(* Logix 5000 project; controller FV vendor 1 type 14 code 217 rev 31.11; software revision 31.00; part 43 of 63 *)
(* tags used below, declared in another part *)
   FV_B100 : INT[255];   // FV FLAGS
   FV_F8 : REAL[256];
   FV_FV10C : PlantItem;   // FV10C
   FV_FV10J : PlantItem;   // FV10J
   FV_FV11C : PlantItem;   // FV11C
   FV_FV11J : PlantItem;   // FV11J
   FV_FV12C : PlantItem;   // FV12C
   FV_FV12J : PlantItem;   // FV12J
   FV_FV13C : PlantItem;   // FV13C
   FV_FV13J : PlantItem;   // FV13J
   FV_FV14C : PlantItem;   // FV14C
   FV_FV14J : PlantItem;   // FV14J
   FV_FV15C : PlantItem;   // FV15C
   FV_FV15J : PlantItem;   // FV15J
   FV_FV16C : PlantItem;   // FV16C
   FV_FV16J : PlantItem;   // FV16J
   FV_FV17C : PlantItem;   // FV17C
   FV_FV17J : PlantItem;   // FV17J
   FV_FV18C : PlantItem;   // FV18C
   FV_FV18J : PlantItem;   // FV18J
   FV_FV19C : PlantItem;   // FV19C
   FV_FV19J : PlantItem;   // FV19J
   FV_FV1C : PlantItem;   // FV1C
   FV_FV1J : PlantItem;   // FV1J
   FV_FV20C : PlantItem;   // FV20C
   FV_FV20J : PlantItem;   // FV20J
   FV_FV21C : PlantItem;   // FV21C
   FV_FV21J : PlantItem;   // FV21J
   FV_FV22C : PlantItem;   // FV22C
   FV_FV22J : PlantItem;   // FV22J
   FV_FV2C : PlantItem;   // FV2C
   FV_FV2J : PlantItem;   // FV2J
   FV_FV3C : PlantItem;   // FV3C
   FV_FV3J : PlantItem;   // FV3J
   FV_FV4C : PlantItem;   // FV4C
   FV_FV4J : PlantItem;   // FV4J
   FV_FV5C : PlantItem;   // FV5C
   FV_FV5J : PlantItem;   // FV5J
   FV_FV6C : PlantItem;   // FV6C
   FV_FV6J : PlantItem;   // FV6J
   FV_FV7C : PlantItem;   // FV7C
   FV_FV7J : PlantItem;   // FV7J
   FV_FV8C : PlantItem;   // FV8C
   FV_FV8J : PlantItem;   // FV8J
   FV_FV9C : PlantItem;   // FV9C
   FV_FV9J : PlantItem;   // FV9J
   FV_N101 : INT[255];   // FV INT Fermentation control integer workspace
   FV_N110 : INT[255];   // FV DATA 0 CURRENT FV DATA
   FV_N111 : INT[50];   // FV1, CURRENT FV DATA
   FV_N112 : INT[50];   // FV2, CURRENT FV DATA
   FV_N113 : INT[50];   // FV3, CURRENT FV DATA
   FV_N114 : INT[50];   // FV4, CURRENT FV DATA
   FV_N115 : INT[50];   // FV5, CURRENT FV DATA
   FV_N116 : INT[50];   // FV6, CURRENT FV DATA
   FV_N117 : INT[50];   // FV7, CURRENT FV DATA
   FV_N118 : INT[50];   // FV8, CURRENT FV DATA
   FV_N119 : INT[50];   // FV9, CURRENT FV DATA
   FV_N12 : INT[255];   // SYS_PARMS System Parameter Fil e
   FV_N120 : INT[50];   // FV10, CURRENT FV DATA
   FV_N121 : INT[50];   // FV11, CURRENT FV DATA
   FV_N122 : INT[50];   // FV12, CURRENT FV DATA
   FV_N123 : INT[50];   // FV13, CURRENT FV DATA
   FV_N124 : INT[50];   // FV14, CURRENT FV DATA
   FV_N125 : INT[50];   // FV15, CURRENT FV DATA
   FV_N126 : INT[50];   // FV16, CURRENT FV DATA
   FV_N127 : INT[50];   // FV17, CURRENT FV DATA
   FV_N128 : INT[50];   // FV18, CURRENT FV DATA
   FV_N129 : INT[50];   // FV19, CURRENT FV DATA
   FV_N130 : INT[50];   // FV20, CURRENT FV DATA
   FV_N131 : INT[50];   // FV21, CURRENT FV DATA
   FV_N132 : INT[50];   // FV22, CURRENT FV DATA
   FV_SFile : INT[255];   // SLC Equivalent System File, So Original Code Can Remain
(* FV_Common, continued *)

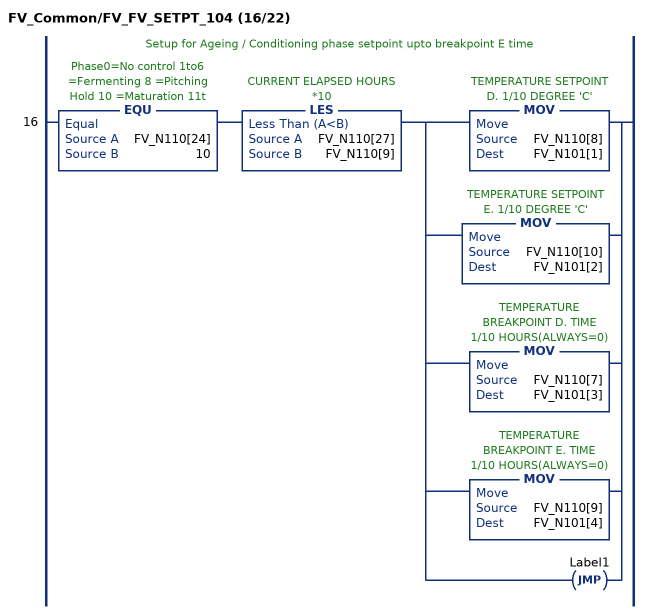
   [picture p920: FV_Common/FV_FV_SETPT_104 rungs 16-16]
   // Setup for Ageing / Conditioning phase setpoint upto breakpoint E time
   16: EQU(FV_N110[24],10)LES(FV_N110[27],FV_N110[9])[MOV(FV_N110[8],FV_N101[1]) ,MOV(FV_N110[10],FV_N101[2]) ,MOV(FV_N110[7],FV_N101[3]) ,MOV(FV_N110[9],FV_N101[4]) ,JMP(Label1) ];
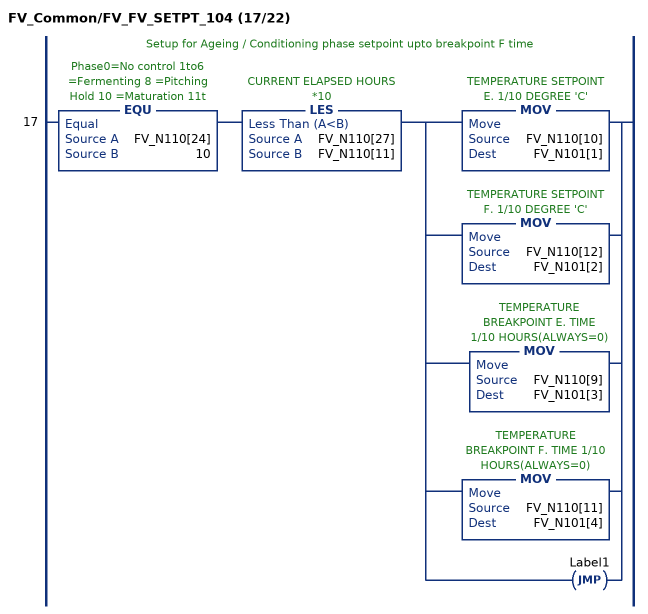
   // Setup for Ageing / Conditioning phase setpoint upto breakpoint F time
   17: EQU(FV_N110[24],10)LES(FV_N110[27],FV_N110[11])[MOV(FV_N110[10],FV_N101[1]) ,MOV(FV_N110[12],FV_N101[2]) ,MOV(FV_N110[9],FV_N101[3]) ,MOV(FV_N110[11],FV_N101[4]) ,JMP(Label1) ];
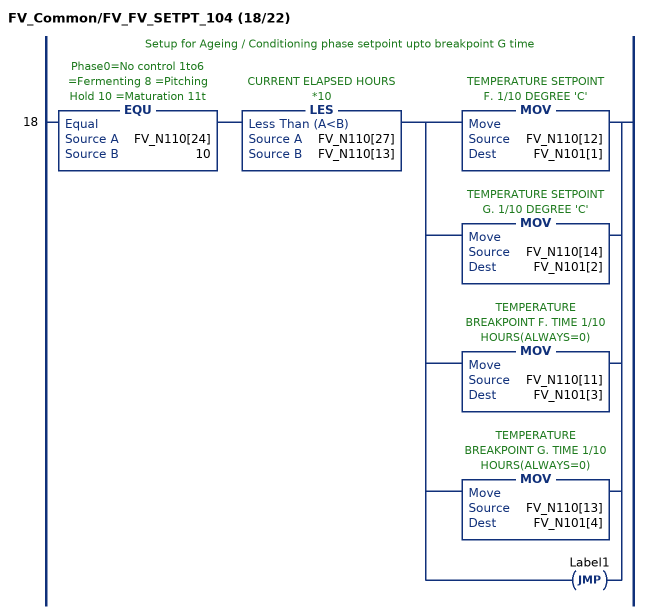
   // Setup for Ageing / Conditioning phase setpoint upto breakpoint G time
   18: EQU(FV_N110[24],10)LES(FV_N110[27],FV_N110[13])[MOV(FV_N110[12],FV_N101[1]) ,MOV(FV_N110[14],FV_N101[2]) ,MOV(FV_N110[11],FV_N101[3]) ,MOV(FV_N110[13],FV_N101[4]) ,JMP(Label1) ];
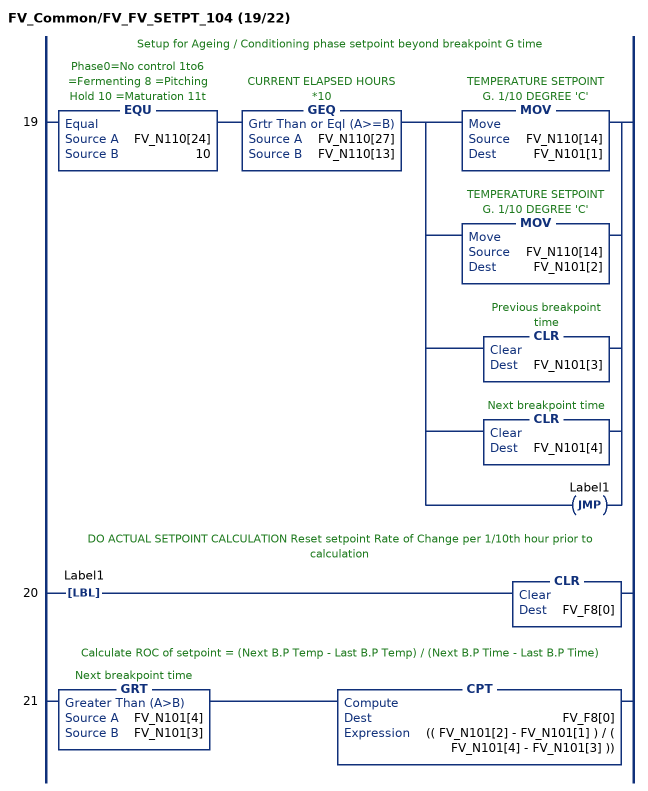
   // Setup for Ageing / Conditioning phase setpoint beyond breakpoint G time
   19: EQU(FV_N110[24],10)GEQ(FV_N110[27],FV_N110[13])[MOV(FV_N110[14],FV_N101[1]) ,MOV(FV_N110[14],FV_N101[2]) ,CLR(FV_N101[3]) ,CLR(FV_N101[4]) ,JMP(Label1) ];
   // DO ACTUAL SETPOINT CALCULATION Reset setpoint Rate of Change per 1/10th hour prior to calculation
   20: LBL(Label1)CLR(FV_F8[0]);
   // Calculate ROC of setpoint = (Next B.P Temp - Last B.P Temp) / (Next B.P Time - Last B.P Time)
   21: GRT(FV_N101[4],FV_N101[3])CPT(FV_F8[0],(( FV_N101[2] - FV_N101[1] ) / ( FV_N101[4] - FV_N101[3] )));
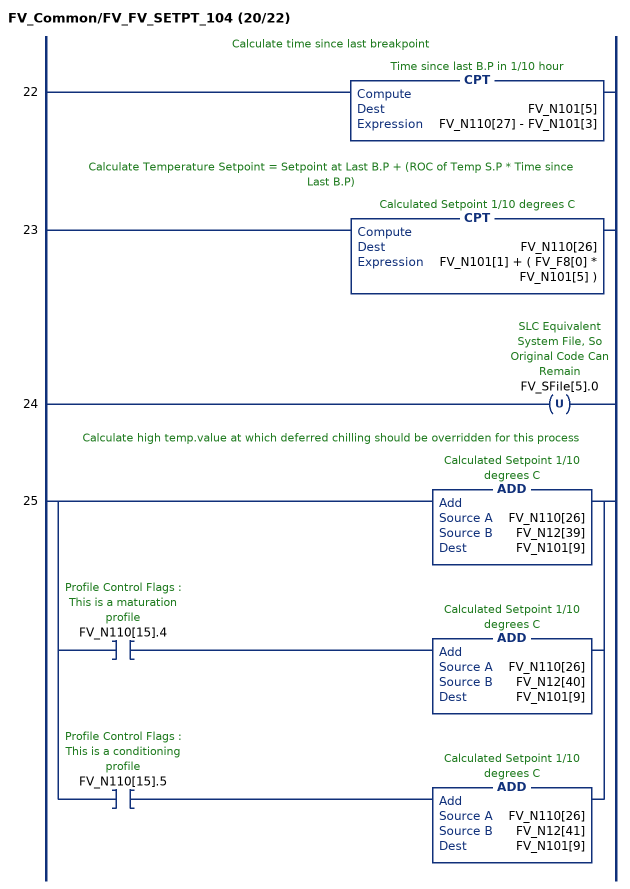
   // Calculate time since last breakpoint
   22: CPT(FV_N101[5],FV_N110[27] - FV_N101[3]);
   // Calculate Temperature Setpoint = Setpoint at Last B.P + (ROC of Temp S.P * Time since Last B.P)
   23: CPT(FV_N110[26],FV_N101[1] + ( FV_F8[0] * FV_N101[5] ));
   24: OTU(FV_SFile[5].0);
   // Calculate high temp.value at which deferred chilling should be overridden for this process
   25: [ADD(FV_N110[26],FV_N12[39],FV_N101[9]) ,XIC(FV_N110[15].4) ADD(FV_N110[26],FV_N12[40],FV_N101[9]) ,XIC(FV_N110[15].5) ADD(FV_N110[26],FV_N12[41],FV_N101[9]) ];
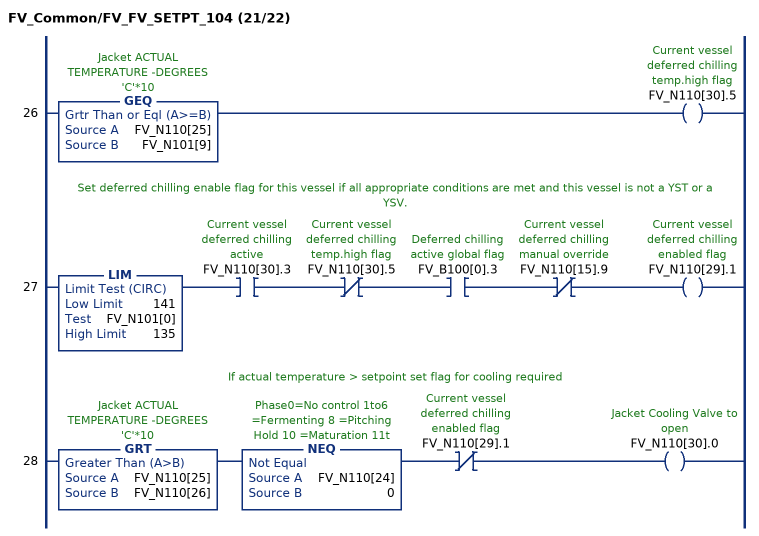
   26: GEQ(FV_N110[25],FV_N101[9])OTE(FV_N110[30].5);
   // Set deferred chilling enable flag for this vessel if all appropriate conditions are met and this vessel is not a YST or a YSV.
   27: LIM(141,FV_N101[0],135)XIC(FV_N110[30].3)XIO(FV_N110[30].5)XIC(FV_B100[0].3)XIO(FV_N110[15].9)OTE(FV_N110[29].1);
   // If actual temperature > setpoint set flag for cooling required
   28: GRT(FV_N110[25],FV_N110[26])NEQ(FV_N110[24],0)XIO(FV_N110[29].1)OTE(FV_N110[30].0);
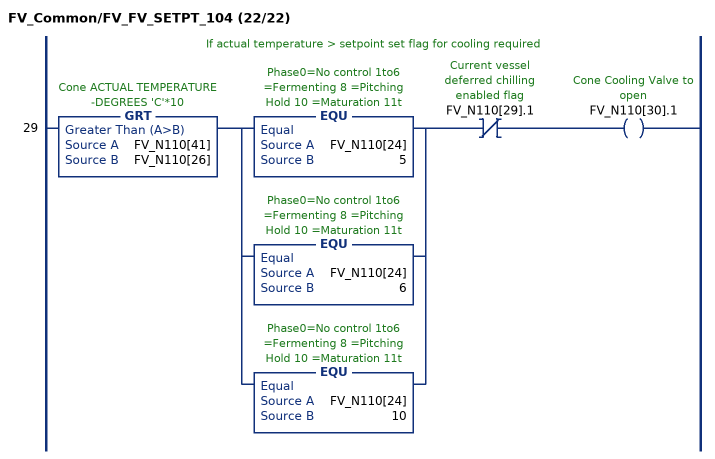
   // If actual temperature > setpoint set flag for cooling required
   29: GRT(FV_N110[41],FV_N110[26])[EQU(FV_N110[24],5) ,EQU(FV_N110[24],6) ,EQU(FV_N110[24],10) ]XIO(FV_N110[29].1)OTE(FV_N110[30].1);
END_ROUTINE

ROUTINE FV_FV_VALVES_105   (* ladder *)
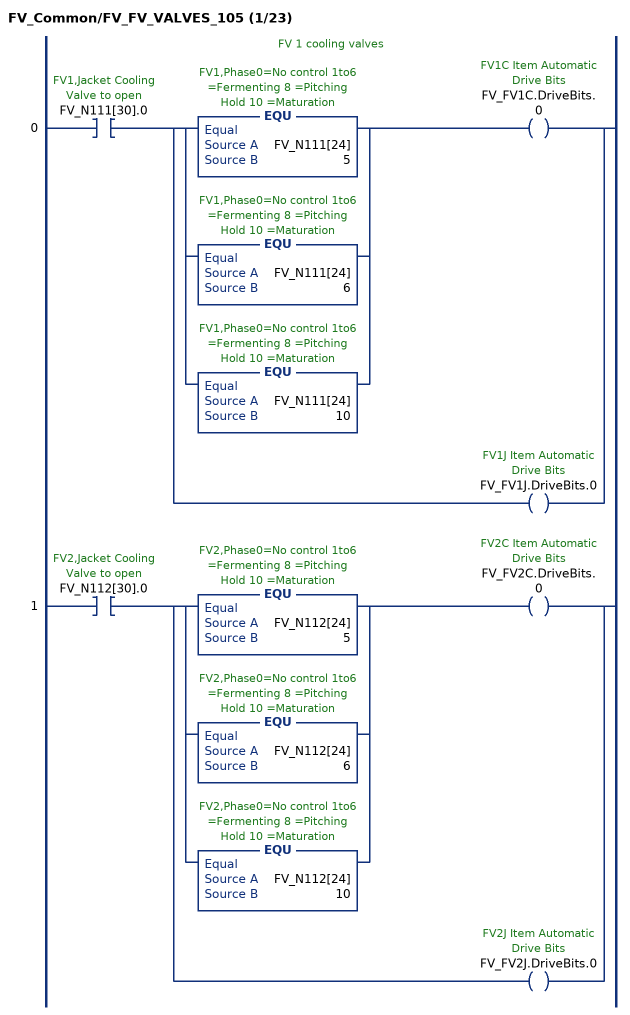
   // FV 1 cooling valves
   0: XIC(FV_N111[30].0)[[EQU(FV_N111[24],5) ,EQU(FV_N111[24],6) ,EQU(FV_N111[24],10) ] OTE(FV_FV1C.DriveBits.0) ,OTE(FV_FV1J.DriveBits.0) ];
   1: XIC(FV_N112[30].0)[[EQU(FV_N112[24],5) ,EQU(FV_N112[24],6) ,EQU(FV_N112[24],10) ] OTE(FV_FV2C.DriveBits.0) ,OTE(FV_FV2J.DriveBits.0) ];
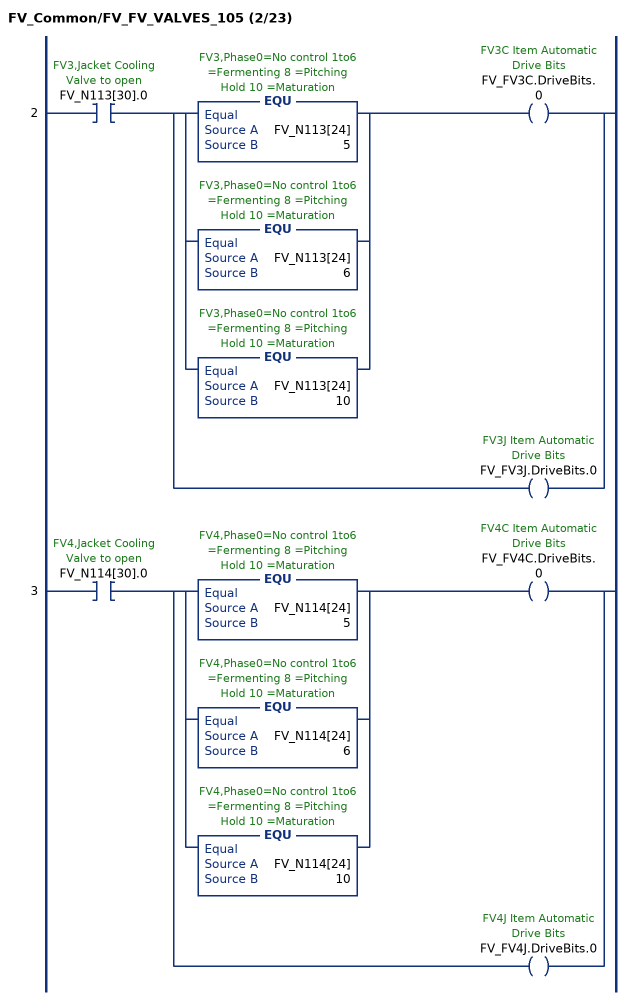
   2: XIC(FV_N113[30].0)[[EQU(FV_N113[24],5) ,EQU(FV_N113[24],6) ,EQU(FV_N113[24],10) ] OTE(FV_FV3C.DriveBits.0) ,OTE(FV_FV3J.DriveBits.0) ];
   3: XIC(FV_N114[30].0)[[EQU(FV_N114[24],5) ,EQU(FV_N114[24],6) ,EQU(FV_N114[24],10) ] OTE(FV_FV4C.DriveBits.0) ,OTE(FV_FV4J.DriveBits.0) ];
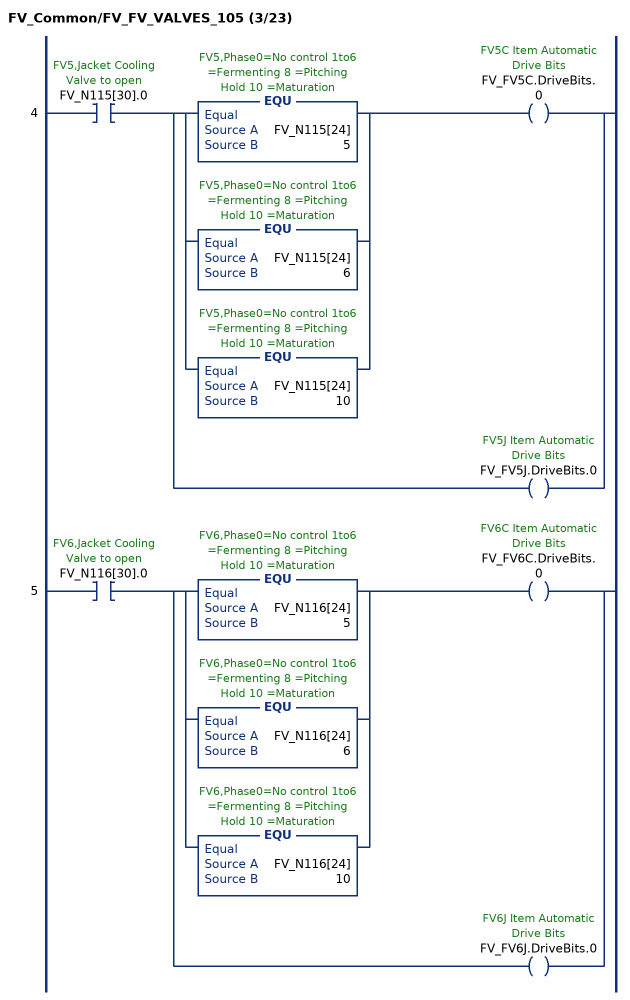
   4: XIC(FV_N115[30].0)[[EQU(FV_N115[24],5) ,EQU(FV_N115[24],6) ,EQU(FV_N115[24],10) ] OTE(FV_FV5C.DriveBits.0) ,OTE(FV_FV5J.DriveBits.0) ];
   5: XIC(FV_N116[30].0)[[EQU(FV_N116[24],5) ,EQU(FV_N116[24],6) ,EQU(FV_N116[24],10) ] OTE(FV_FV6C.DriveBits.0) ,OTE(FV_FV6J.DriveBits.0) ];
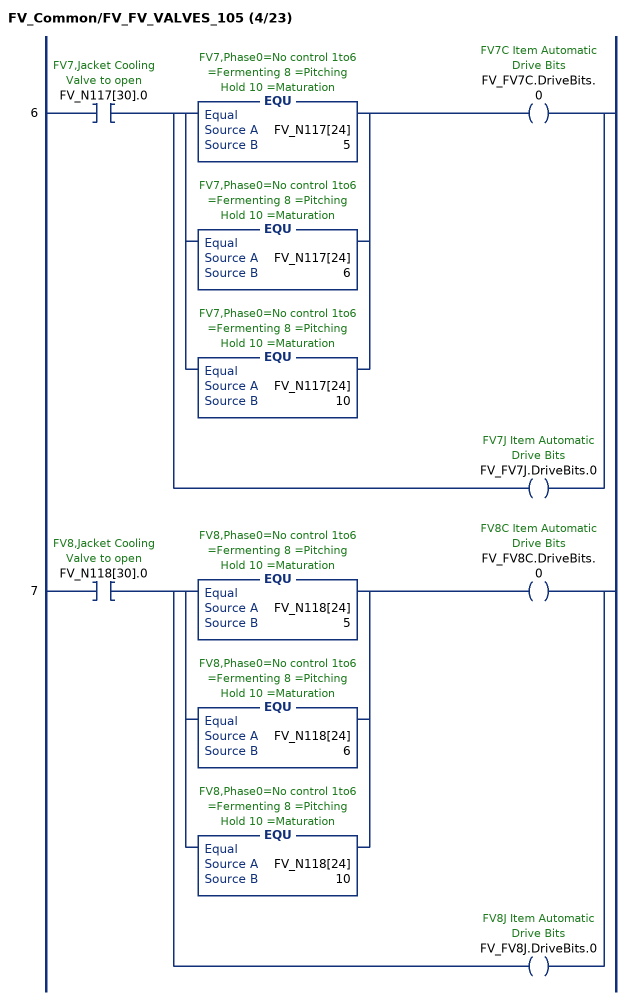
   6: XIC(FV_N117[30].0)[[EQU(FV_N117[24],5) ,EQU(FV_N117[24],6) ,EQU(FV_N117[24],10) ] OTE(FV_FV7C.DriveBits.0) ,OTE(FV_FV7J.DriveBits.0) ];
   7: XIC(FV_N118[30].0)[[EQU(FV_N118[24],5) ,EQU(FV_N118[24],6) ,EQU(FV_N118[24],10) ] OTE(FV_FV8C.DriveBits.0) ,OTE(FV_FV8J.DriveBits.0) ];
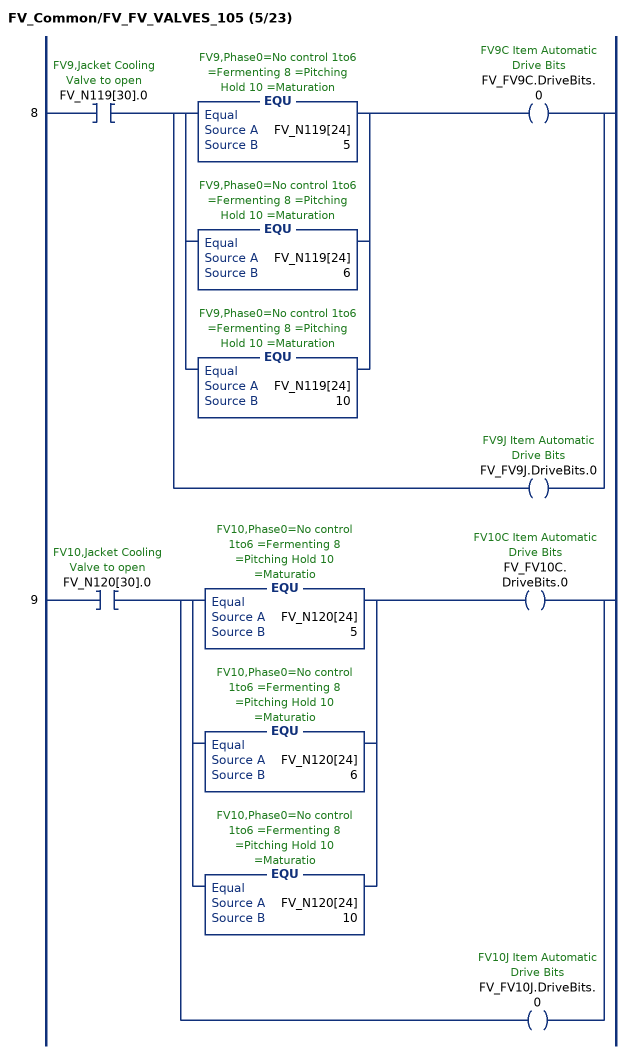
   8: XIC(FV_N119[30].0)[[EQU(FV_N119[24],5) ,EQU(FV_N119[24],6) ,EQU(FV_N119[24],10) ] OTE(FV_FV9C.DriveBits.0) ,OTE(FV_FV9J.DriveBits.0) ];
   9: XIC(FV_N120[30].0)[[EQU(FV_N120[24],5) ,EQU(FV_N120[24],6) ,EQU(FV_N120[24],10) ] OTE(FV_FV10C.DriveBits.0) ,OTE(FV_FV10J.DriveBits.0) ];
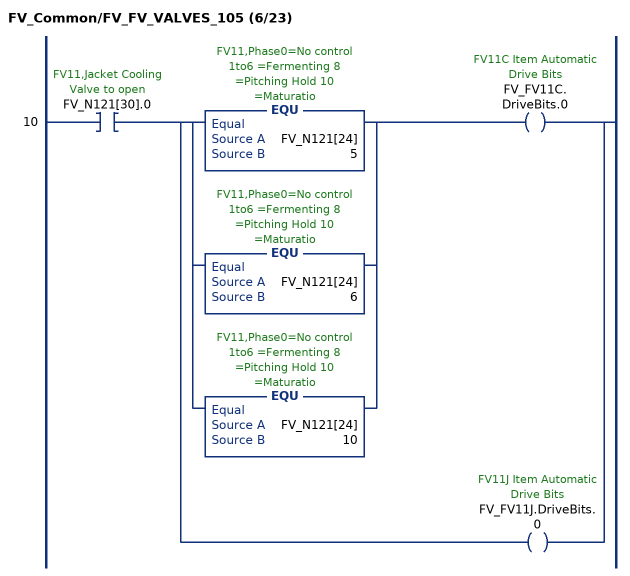
   10: XIC(FV_N121[30].0)[[EQU(FV_N121[24],5) ,EQU(FV_N121[24],6) ,EQU(FV_N121[24],10) ] OTE(FV_FV11C.DriveBits.0) ,OTE(FV_FV11J.DriveBits.0) ];
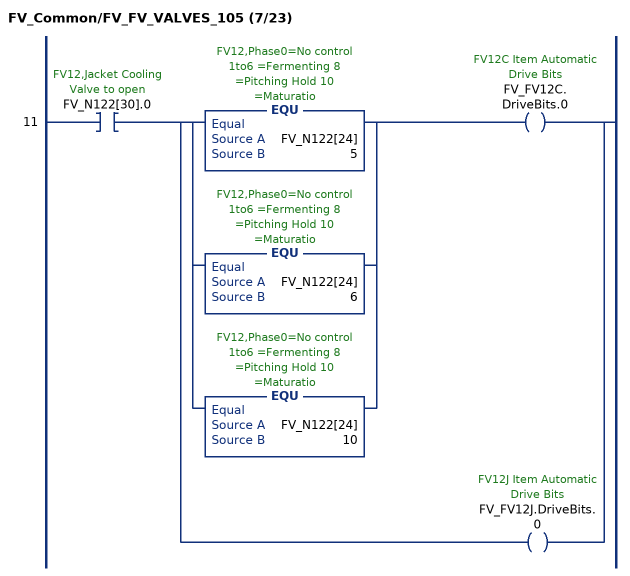
   11: XIC(FV_N122[30].0)[[EQU(FV_N122[24],5) ,EQU(FV_N122[24],6) ,EQU(FV_N122[24],10) ] OTE(FV_FV12C.DriveBits.0) ,OTE(FV_FV12J.DriveBits.0) ];
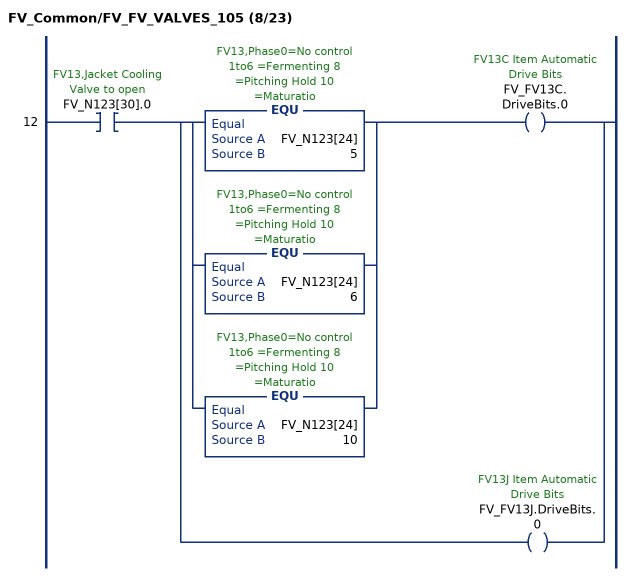
   12: XIC(FV_N123[30].0)[[EQU(FV_N123[24],5) ,EQU(FV_N123[24],6) ,EQU(FV_N123[24],10) ] OTE(FV_FV13C.DriveBits.0) ,OTE(FV_FV13J.DriveBits.0) ];
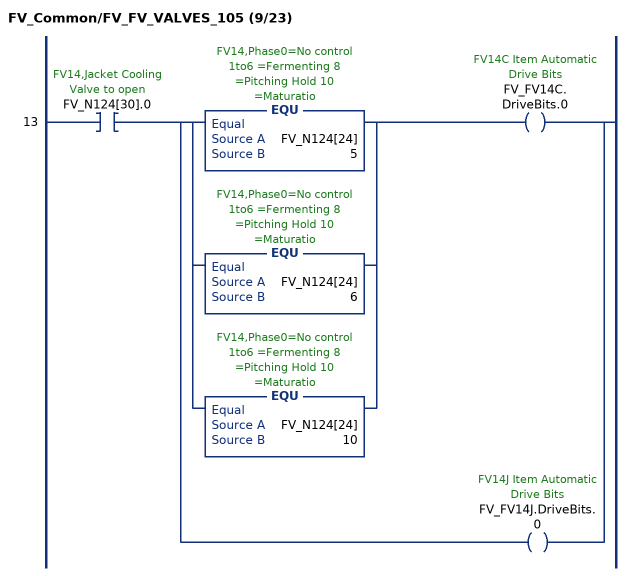
   13: XIC(FV_N124[30].0)[[EQU(FV_N124[24],5) ,EQU(FV_N124[24],6) ,EQU(FV_N124[24],10) ] OTE(FV_FV14C.DriveBits.0) ,OTE(FV_FV14J.DriveBits.0) ];
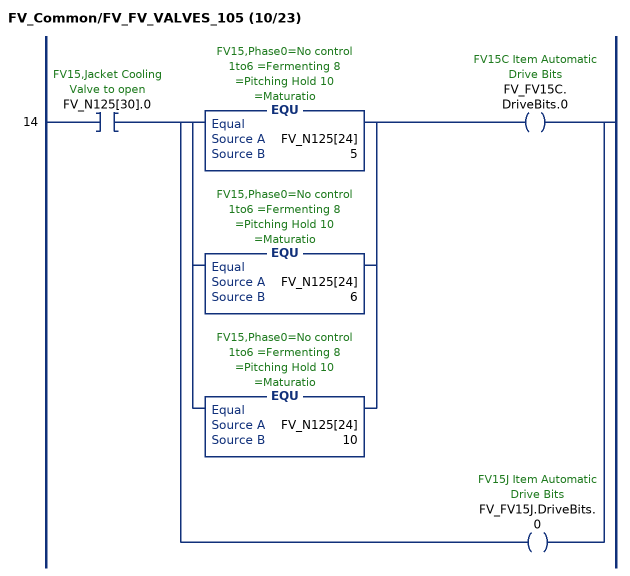
   14: XIC(FV_N125[30].0)[[EQU(FV_N125[24],5) ,EQU(FV_N125[24],6) ,EQU(FV_N125[24],10) ] OTE(FV_FV15C.DriveBits.0) ,OTE(FV_FV15J.DriveBits.0) ];
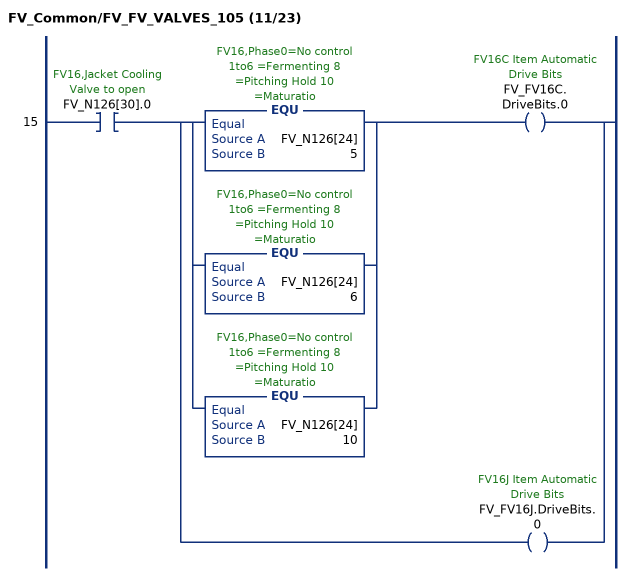
   15: XIC(FV_N126[30].0)[[EQU(FV_N126[24],5) ,EQU(FV_N126[24],6) ,EQU(FV_N126[24],10) ] OTE(FV_FV16C.DriveBits.0) ,OTE(FV_FV16J.DriveBits.0) ];
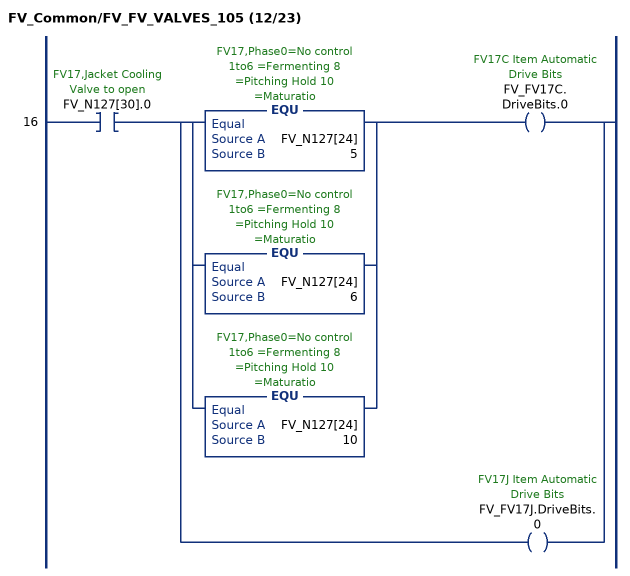
   16: XIC(FV_N127[30].0)[[EQU(FV_N127[24],5) ,EQU(FV_N127[24],6) ,EQU(FV_N127[24],10) ] OTE(FV_FV17C.DriveBits.0) ,OTE(FV_FV17J.DriveBits.0) ];
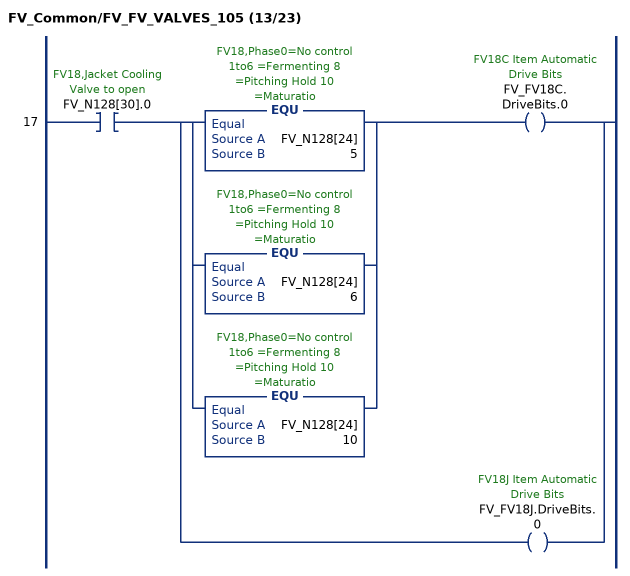
   17: XIC(FV_N128[30].0)[[EQU(FV_N128[24],5) ,EQU(FV_N128[24],6) ,EQU(FV_N128[24],10) ] OTE(FV_FV18C.DriveBits.0) ,OTE(FV_FV18J.DriveBits.0) ];
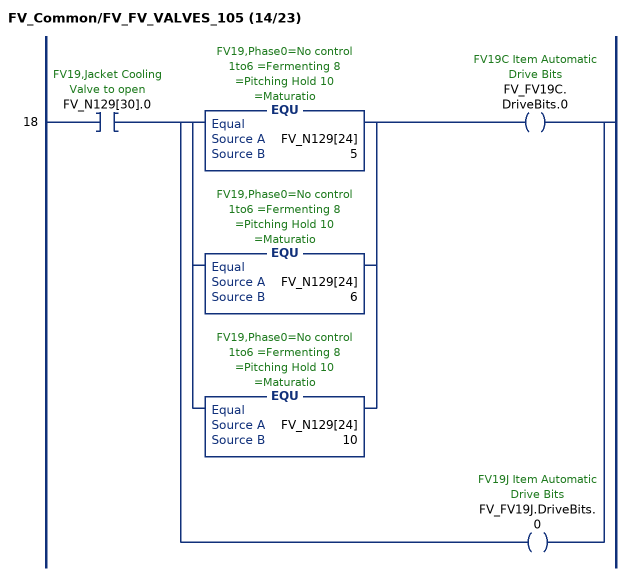
   18: XIC(FV_N129[30].0)[[EQU(FV_N129[24],5) ,EQU(FV_N129[24],6) ,EQU(FV_N129[24],10) ] OTE(FV_FV19C.DriveBits.0) ,OTE(FV_FV19J.DriveBits.0) ];
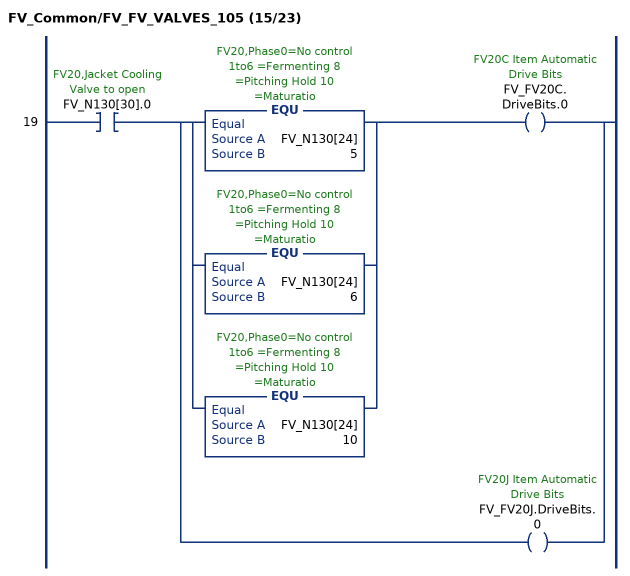
   19: XIC(FV_N130[30].0)[[EQU(FV_N130[24],5) ,EQU(FV_N130[24],6) ,EQU(FV_N130[24],10) ] OTE(FV_FV20C.DriveBits.0) ,OTE(FV_FV20J.DriveBits.0) ];
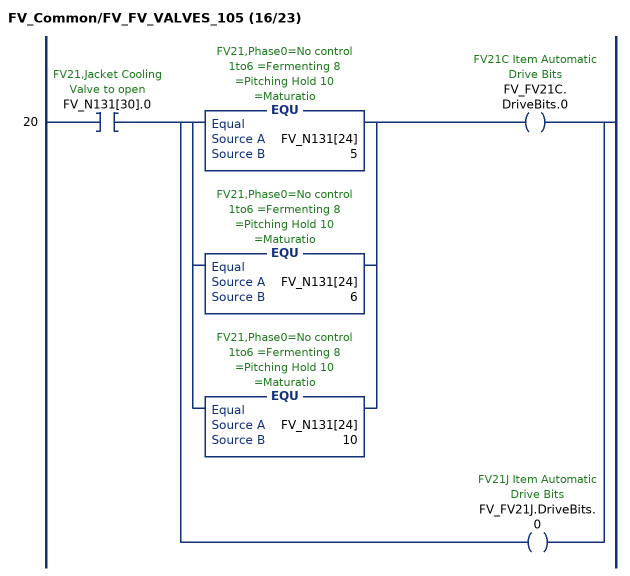
   20: XIC(FV_N131[30].0)[[EQU(FV_N131[24],5) ,EQU(FV_N131[24],6) ,EQU(FV_N131[24],10) ] OTE(FV_FV21C.DriveBits.0) ,OTE(FV_FV21J.DriveBits.0) ];
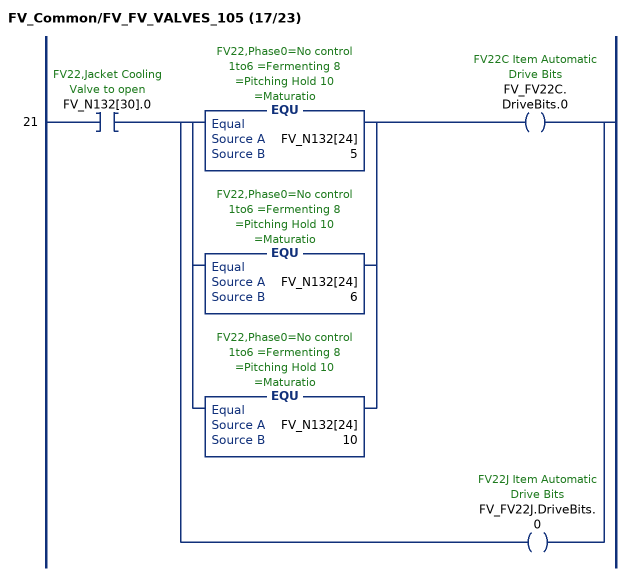
   21: XIC(FV_N132[30].0)[[EQU(FV_N132[24],5) ,EQU(FV_N132[24],6) ,EQU(FV_N132[24],10) ] OTE(FV_FV22C.DriveBits.0) ,OTE(FV_FV22J.DriveBits.0) ];
